'~Spare FB1[273].28'; 8765 '~Spare FB1[273].29'; 8766 '~Spare FB1[273].30'; 8767 '~Spare FB1[273].31'; 8768 '~Spare FB1[274].0'; 8769 '~Spare FB1[274].1'; 8770 '~Spare FB1[274].2'; 8771 '~Spare FB1[274].3'; 8772 '~Spare FB1[274].4'; 8773 '~Spare FB1[274].5'; 8774 '~Spare FB1[274].6'; 8775 '~Spare FB1[274].7'; 8776 '~Spare FB1[274].8'; 8777 '~Spare FB1[274].9'; 8778 '~Spare FB1[274].10'; 8779 '~Spare FB1[274].11'; 8780 '~Spare FB1[274].12'; 8781 '~Spare FB1[274].13'; 8782 '~Spare FB1[274].14'; 8783 '~Spare FB1[274].15'; 8784 '~Spare FB1[274].16'; 8785 '~Spare FB1[274].17'; 8786 '~Spare FB1[274].18'; 8787 '~Spare FB1[274].19'; 8788 '~Spare FB1[274].20'; 8789 '~Spare FB1[274].21'; 8790 '~Spare FB1[274].22'; 8791 '~Spare FB1[274].23'; 8792 '~Spare FB1[274].24'; 8793 '~Spare FB1[274].25'; 8794 '~Spare FB1[274].26'; 8795 '~Spare FB1[274].27'; 8796 '~Spare FB1[274].28'; 8797 '~Spare FB1[274].29'; 8798 '~Spare FB1[274].30'; 8799 '~Spare FB1[274].31'; 8800 '~Spare FB1[275].0'; 8801 '~Spare FB1[275].1'; 8802 '~Spare FB1[275].2'; 8803 '~Spare FB1[275].3'; 8804 '~Spare FB1[275].4'; 8805 '~Spare FB1[275].5'; 8806 '~Spare FB1[275].6'; 8807 '~Spare FB1[275].7'; 8808 '~Spare FB1[275].8'; 8809 '~Spare FB1[275].9'; 8810 '~Spare FB1[275].10'; 8811 '~Spare FB1[275].11'; 8812 '~Spare FB1[275].12'; 8813 '~Spare FB1[275].13'; 8814 '~Spare FB1[275].14'; 8815 '~Spare FB1[275].15'; 8816 '~Spare FB1[275].16'; 8817 '~Spare FB1[275].17'; 8818 '~Spare FB1[275].18'; 8819 '~Spare FB1[275].19'; 8820 '~Spare FB1[275].20'; 8821 '~Spare FB1[275].21'; 8822 '~Spare FB1[275].22'; 8823 '~Spare FB1[275].23'; 8824 '~Spare FB1[275].24'; 8825 '~Spare FB1[275].25'; 8826 '~Spare FB1[275].26'; 8827 '~Spare FB1[275].27'; 8828 '~Spare FB1[275].28'; 8829 '~Spare FB1[275].29'; 8830 '~Spare FB1[275].30'; 8831 '~Spare FB1[275].31'; 8832 '~S001R05CN.I.RbtCtrlFlt - Control Fault FB1[276].0'; 8833 '~S001R05CN.I.CollDetect - Collision Detect FB1[276].1'; 8834 '~S001R05CN.Ix.RbtPromptBox - View Prompt Box at Teach Pendant FB1[276].2'; 8835 '~Spare FB1[276].3'; 8836 '~Spare FB1[276].4'; 8837 '~Spare FB1[276].5'; 8838 '~Spare FB1[276].6'; 8839 '~Spare FB1[276].7'; 8840 '~Spare FB1[276].8'; 8841 '~Spare FB1[276].9'; 8842 '~Spare FB1[276].10'; 8843 '~S001R05CN.I.Wc1WldFlt -Weld Controller 1 Weld Fault FB1[276].11'; 8844 '~S001R05CN.I.Wc1Flt - Weld Timer Flt - Depress Man Weld To Continue FB1[276].12'; 8845 '~S001R05CN.I.Wc1SGunFlt - Weld Controller 1 Servo Gun Fault FB1[276].13'; 8846 '~S001R05CN.I.Wc1SGunMtrTempFlt - Cntrl 1 Servo Gun Motor Over Temp FB1[276].14'; 8847 '~S001R05CN.I.Td1MtrFlt - Tip Dress 1 Motor Fault FB1[276].15'; 8848 '~S001R05CN.I.WC1XfmrTempFlt - Weld Cntrl 1 Transformer Over Temp FB1[276].16'; 8849 '~S001R05CN.I.AutoTipChng1Flt - Auto Tip Changer 1 Fault FB1[276].17'; 8850 '~S001R05CN.I.Slr1NotReady - Seal Controller 1 Not Ready FB1[276].18'; 8851 '~S001R05CN.I.Slr1MajorFlt - Seal Controller 1 Major Fault FB1[276].19'; 8852 '~S001R05CN.I.Slr1VolNotOk - Seal Controller 1 Volume Not Ok Fault FB1[276].20'; 8853 '~S001R05CN.I.Slr1PurgeFlt - Seal Controller 1 Purge Fault FB1[276].21'; 8854 '~S001R05CN.I.Slr1DoserNot Filled - Seal Cntrl 1 Doser Not Filled FB1[276].22'; 8855 '~S001R05CN.I.Slr1No2ClnMxr - Seal Cntrl1 No 2C In Mixer Fault FB1[276].23'; 8856 '~S001R05CN.I.Slr1NzlBroken - Seal Controller 1 Nozzle Broken Fault FB1[276].24'; 8857 '~S001R05CN.I.Slr1NozzleChgReq - Seal Cntrl1 Nozzle Change Reqd FB1[276].25'; 8858 '~S001R05CN.I.Slr1CycleInterrupted - Seal Cntrl1 Cycle Interrupted FB1[276].26'; 8859 '~S001R05CN.I.Stdw1Flt - Stud Weld 1 Weld Fault FB1[276].27'; 8860 '~S001R05CN.I.Stdw1DlyExcdd - Stud Weld 1 Time Delay Exceeded Flt FB1[276].28'; 8861 '~S001R05CN.I.Stdw1Maint Reqd - Stud Weld 1 Maintenance Required FB1[276].29'; 8862 '~S001R05CN.I.Stdw1Reject - Stud Weld 1 art Reject Fault FB1[276].30'; 8863 '~S001R05CN.I.Rvt1Flt - Rivet Controller 1 Fault FB1[276].31'; 8864 '~S001R05CN.I.Rvt1DlyExcdd - Rivet Cntrl 1 Time Delay Exceeded Flt FB1[277].0'; 8865 '~S001R05CN.I.AutoPulledTipByp1 - Auto Pulled Tip Bypass 1 FB1[277].1'; 8866 '~S001R05CN.I.StdWld1EquipmentFlt - Stud Weld 1 Equipment Fault FB1[277].2'; 8867 '~S001R05CN.I.StdWld1BrcktNotPresent - Stud Weld 1 Bracket Not Pres FB1[277].3'; 8868 '~S001R05CN.I.PierceFlt - Pierce Fault FB1[277].4'; 8869 '~S001R05CN.I.NoVisionMeasErr - Vision System Measurement Error FB1[277].5'; 8870 '~S001R05CN.I.VisionSysCalErr - Vision System Calibration Fault FB1[277].6'; 8871 '~S001R05CN.I.VisionSysErr - Vision System Error FB1[277].7'; 8872 '~S001R05CN.I.RackOutOfTolerance - Vision Sys Rack Out Of Tolerance FB1[277].8'; 8873 '~S001R05CN.Ix.TorqFlt - Torque Not Ok FB1[277].9'; 8874 '~S001R05CN.Ix.MwFlt - Mig Weld Controller Fault FB1[277].10'; 8875 '~S001R05CN.Ix.MwWireStuckFlt - Mig Welder Wire Stuck FB1[277].11'; 8876 '~S001R05CN.Ix.MwWldFlt - Mig Welder Bad Bronze Weld Indicator Flt FB1[277].12'; 8877 '~S001R05CN.I.O.TipChngReqd1 - Weld Cntrl 1 Tip Change Required FB1[277].13'; 8878 '~S001R05CN.I.M.NutDetectFlt1 - Nut Welder 1 Nut Detection Fault FB1[277].14'; 8879 '~S001R05CN.I.M.NutProjFlt1 - Nut Welder 1 Weld Not In Tolerance FB1[277].15'; 8880 '~S001R05CN.M.WrongRivetAtNose - Remove Wrong Rivet At Nose FB1[277].16'; 8881 '~S001R05CN.Ix.MwWldLimitErr - Mig Welder CurrentVoltage Out of Tolerance FB1[277].17'; 8882 '~S001R05CN.Ix.MigRdy Mig Welder Not Ready FB1[277].18'; 8883 '~Spare FB1[277].19'; 8884 '~Spare FB1[277].20'; 8885 '~S001R05CN.I.Wc2WldFlt -Weld Controller 2 Weld Fault FB1[277].21'; 8886 '~S001R05CN.I.Wc2Flt - Weld Timer Flt - Depress Man Weld To Continue FB1[277].22'; 8887 '~S001R05CN.I.Wc2SGunFlt - Weld Controller 2 Servo Gun Fault FB1[277].23'; 8888 '~S001R05CN.I.Wc2SGunMtrTempFlt - Cntrl 2 Servo Gun Motor Over Temp FB1[277].24'; 8889 '~S001R05CN.I.Td2MtrFlt - Tip Dress 2 Motor Fault FB1[277].25'; 8890 '~S001R05CN.I.WC2XfmrTempFlt - Weld Cntrl 2 Transformer Over Temp FB1[277].26'; 8891 '~S001R05CN.I.AutoTipChng2Flt - Auto Tip Changer 2 Fault FB1[277].27'; 8892 '~S001R05CN.I.Slr2NotReady - Seal Controller 2 Not Ready FB1[277].28'; 8893 '~S001R05CN.I.Slr2MajorFlt - Seal Controller 2 Major Fault FB1[277].29'; 8894 '~S001R05CN.I.Slr2VolNotOk - Seal Controller 2 Volume Not Ok Fault FB1[277].30'; 8895 '~S001R05CN.I.Slr2PurgeFlt - Seal Controller 2 Purge Fault FB1[277].31'; 8896 '~S001R05CN.I.Slr2DoserNot Filled - Seal Cntrl 2 Doser Not Filled FB1[278].0'; 8897 '~S001R05CN.I.Slr2No2ClnMxr - Seal Cntrl2 No 2C In Mixer Fault FB1[278].1'; 8898 '~S001R05CN.I.Slr2NzlBroken - Seal Controller 2 Nozzle Broken Fault FB1[278].2'; 8899 '~S001R05CN.I.Slr2NozzleChgReq - Seal Cntrl2 Nozzle Change Reqd FB1[278].3'; 8900 '~S001R05CN.I.Slr2CycleInterrupted - Seal Cntrl2 Cycle Interrupted FB1[278].4'; 8901 '~S001R05CN.I.Stdw2Flt - Stud Weld 2 Weld Fault FB1[278].5'; 8902 '~S001R05CN.I.Stdw2DlyExcdd - Stud Weld 2 Time Delay Exceeded Flt FB1[278].6'; 8903 '~S001R05CN.I.Stdw2Maint Reqd - Stud Weld 2 Maintenance Required FB1[278].7'; 8904 '~S001R05CN.I.Stdw2Reject - Stud Weld 2 art Reject Fault FB1[278].8'; 8905 '~S001R05CN.I.Rvt2Flt - Rivet Controller 2 Fault FB1[278].9'; 8906 '~S001R05CN.I.Rvt2DlyExcdd - Rivet Cntrl 2 Time Delay Exceeded Flt FB1[278].10'; 8907 '~S001R05CN.I.AutoPulledTipByp2 - Auto Pulled Tip Bypass 2 FB1[278].11'; 8908 '~S001R05CN.I.StdWld2EquipmentFlt - Stud Weld 2 Equipment Fault FB1[278].12'; 8909 '~S001R05CN.I.StdWld2BrcktNotPresent - Stud Weld 2 Bracket Not Pres FB1[278].13'; 8910 '~S001R05CN.Ix.LsrWldMntrFlt - Seam Geometry/Laser Weld Monitor Flt FB1[278].14'; 8911 '~S001R05CN.Ix.LsrHeadFlt - Laser Head Fault FB1[278].15'; 8912 '~S001R05CN.Ix.LsrGlsFlt - Glass Fault FB1[278].16'; 8913 '~S001R05CN.Ix.LsrWhlFlt - Pressure Wheel Not In Range Fault FB1[278].17'; 8914 '~S001R05CN.Ix.LsrGeoFlt - Seam Geometry/Laser Bad Process Geo Flt FB1[278].18'; 8915 '~S001R05CN.Ix.LsrHdCollFlt - Laser Head Collision Fault FB1[278].19'; 8916 '~S001R05CN.Ix.LsrHdSysFlt - Laser Head System Fault FB1[278].20'; 8917 '~S001R05CN.Ix.LsrHdFar - Laser Head Far Fault FB1[278].21'; 8918 '~S001R05CN.Ix.LsrHdSftCollFlt - Laser Head Software Collision Flt FB1[278].22'; 8919 '~S001R05CN.I.O.TipChngReqd2 - Weld Cntrl 2 Tip Change Required FB1[278].23'; 8920 '~S001R05CN.I.M.NutDetectFlt2 - Nut Welder 2 Nut Detection Fault FB1[278].24'; 8921 '~S001R05CN.I.M.NutProjFlt2 - Nut Welder 2 Weld Not In Tolerance FB1[278].25'; 8922 '~S001R05CN.I.TCWrongToolInStand - Tool Changer Wrong Tool In Stand FB1[278].26'; 8923 '~Spare FB1[278].27'; 8924 '~Spare FB1[278].28'; 8925 '~Spare FB1[278].29'; 8926 '~Spare FB1[278].30'; 8927 '~Spare FB1[278].31'; 8928 '~S001R05CN.I.VisionCommOK - Vision System Comm Fault FB1[279].0'; 8929 '~S001R05CN.I.OutOfTolerance - Vision System Out Of Tolerance FB1[279].1'; 8930 '~S001R05CN.I.MeasureReject - Vision System Measure Reject FB1[279].2'; 8931 '~S001R05CN.I.VisionSysCalibrationFlt - Vision System Calibration Flt FB1[279].3'; 8932 '~S001R05CN.I.VisionSysFlt - Vision System Flt FB1[279].4'; 8933 '~Spare FB1[279].5'; 8934 '~Spare FB1[279].6'; 8935 '~Spare FB1[279].7'; 8936 '~Spare FB1[279].8'; 8937 '~Spare FB1[279].9'; 8938 '~Spare FB1[279].10'; 8939 '~Spare FB1[279].11'; 8940 '~Spare FB1[279].12'; 8941 '~Spare FB1[279].13'; 8942 '~Spare FB1[279].14'; 8943 '~Spare FB1[279].15'; 8944 '~Spare FB1[279].16'; 8945 '~Spare FB1[279].17'; 8946 '~S001R05CN.M.InteruptCyc - Laser Cyc Interupt Cut Wire And Reject Car FB1[279].18'; 8947 '~S001R05CN.M.SuspectPart Inspect Vehicle And Accept Or Reject FB1[279].19'; 8948 '~S001R05 Power Meter High Power Fault Detected FB1[279].20'; 8949 '~S001R05 Power Meter Low Power Fault Detected FB1[279].21'; 8950 '~Spare FB1[279].22'; 8951 '~Spare FB1[279].23'; 8952 '~Spare FB1[279].24'; 8953 '~Spare FB1[279].25'; 8954 '~Spare FB1[279].26'; 8955 '~Spare FB1[279].27'; 8956 '~Spare FB1[279].28'; 8957 '~Spare FB1[279].29'; 8958 '~Spare FB1[279].30'; 8959 '~Spare FB1[279].31'; 8960 '~Spare FB1[280].0'; 8961 '~Spare FB1[280].1'; 8962 '~Spare FB1[280].2'; 8963 '~Spare FB1[280].3'; 8964 '~Spare FB1[280].4'; 8965 '~Spare FB1[280].5'; 8966 '~Spare FB1[280].6'; 8967 '~Spare FB1[280].7'; 8968 '~Spare FB1[280].8'; 8969 '~Spare FB1[280].9'; 8970 '~Spare FB1[280].10'; 8971 '~Spare FB1[280].11'; 8972 '~Spare FB1[280].12'; 8973 '~Spare FB1[280].13'; 8974 '~Spare FB1[280].14'; 8975 '~Spare FB1[280].15'; 8976 '~Spare FB1[280].16'; 8977 '~Spare FB1[280].17'; 8978 '~Spare FB1[280].18'; 8979 '~Spare FB1[280].19'; 8980 '~Spare FB1[280].20'; 8981 '~Spare FB1[280].21'; 8982 '~Spare FB1[280].22'; 8983 '~Spare FB1[280].23'; 8984 '~Spare FB1[280].24'; 8985 '~Spare FB1[280].25'; 8986 '~Spare FB1[280].26'; 8987 '~Spare FB1[280].27'; 8988 '~Spare FB1[280].28'; 8989 '~Spare FB1[280].29'; 8990 '~Spare FB1[280].30'; 8991 '~Spare FB1[280].31'; 8992 '~Spare FB1[281].0'; 8993 '~Spare FB1[281].1'; 8994 '~Spare FB1[281].2'; 8995 '~Spare FB1[281].3'; 8996 '~Spare FB1[281].4'; 8997 '~Spare FB1[281].5'; 8998 '~Spare FB1[281].6'; 8999 '~Spare FB1[281].7'; 9000 '~Spare FB1[281].8'; 9001 '~Spare FB1[281].9'; 9002 '~Spare FB1[281].10'; 9003 '~Spare FB1[281].11'; 9004 '~Spare FB1[281].12'; 9005 '~Spare FB1[281].13'; 9006 '~Spare FB1[281].14'; 9007 '~Spare FB1[281].15'; 9008 '~Spare FB1[281].16'; 9009 '~Spare FB1[281].17'; 9010 '~Spare FB1[281].18'; 9011 '~Spare FB1[281].19'; 9012 '~Spare FB1[281].20'; 9013 '~Spare FB1[281].21'; 9014 '~Spare FB1[281].22'; 9015 '~Spare FB1[281].23'; 9016 '~Spare FB1[281].24'; 9017 '~Spare FB1[281].25'; 9018 '~Spare FB1[281].26'; 9019 '~Spare FB1[281].27'; 9020 '~Spare FB1[281].28'; 9021 '~Spare FB1[281].29'; 9022 '~Spare FB1[281].30'; 9023 '~Spare FB1[281].31'; 9024 '~Spare FB1[282].0'; 9025 '~Spare FB1[282].1'; 9026 '~Spare FB1[282].2'; 9027 '~Spare FB1[282].3'; 9028 '~Spare FB1[282].4'; 9029 '~Spare FB1[282].5'; 9030 '~Spare FB1[282].6'; 9031 '~Spare FB1[282].7'; 9032 '~Spare FB1[282].8'; 9033 '~Spare FB1[282].9'; 9034 '~Spare FB1[282].10'; 9035 '~Spare FB1[282].11'; 9036 '~Spare FB1[282].12'; 9037 '~Spare FB1[282].13'; 9038 '~Spare FB1[282].14'; 9039 '~Spare FB1[282].15'; 9040 '~Spare FB1[282].16'; 9041 '~Spare FB1[282].17'; 9042 '~Spare FB1[282].18'; 9043 '~Spare FB1[282].19'; 9044 '~Spare FB1[282].20'; 9045 '~Spare FB1[282].21'; 9046 '~Spare FB1[282].22'; 9047 '~Spare FB1[282].23'; 9048 '~Spare FB1[282].24'; 9049 '~Spare FB1[282].25'; 9050 '~Spare FB1[282].26'; 9051 '~Spare FB1[282].27'; 9052 '~Spare FB1[282].28'; 9053 '~Spare FB1[282].29'; 9054 '~Spare FB1[282].30'; 9055 '~Spare FB1[282].31'; 9056 '~Spare FB1[283].0'; 9057 '~Spare FB1[283].1'; 9058 '~Spare FB1[283].2'; 9059 '~Spare FB1[283].3'; 9060 '~Spare FB1[283].4'; 9061 '~Spare FB1[283].5'; 9062 '~Spare FB1[283].6'; 9063 '~Spare FB1[283].7'; 9064 '~Spare FB1[283].8'; 9065 '~Spare FB1[283].9'; 9066 '~Spare FB1[283].10'; 9067 '~Spare FB1[283].11'; 9068 '~Spare FB1[283].12'; 9069 '~Spare FB1[283].13'; 9070 '~Spare FB1[283].14'; 9071 '~Spare FB1[283].15'; 9072 '~Spare FB1[283].16'; 9073 '~Spare FB1[283].17'; 9074 '~Spare FB1[283].18'; 9075 '~Spare FB1[283].19'; 9076 '~Spare FB1[283].20'; 9077 '~Spare FB1[283].21'; 9078 '~Spare FB1[283].22'; 9079 '~Spare FB1[283].23'; 9080 '~Spare FB1[283].24'; 9081 '~Spare FB1[283].25'; 9082 '~Spare FB1[283].26'; 9083 '~Spare FB1[283].27'; 9084 '~Spare FB1[283].28'; 9085 '~Spare FB1[283].29'; 9086 '~Spare FB1[283].30'; 9087 '~Spare FB1[283].31'; 9088 '~S001R06CN.I.RbtCtrlFlt - Control Fault FB1[284].0'; 9089 '~S001R06CN.I.CollDetect - Collision Detect FB1[284].1'; 9090 '~S001R06CN.Ix.RbtPromptBox - View Prompt Box at Teach Pendant FB1[284].2'; 9091 '~Spare FB1[284].3'; 9092 '~Spare FB1[284].4'; 9093 '~Spare FB1[284].5'; 9094 '~Spare FB1[284].6'; 9095 '~Spare FB1[284].7'; 9096 '~Spare FB1[284].8'; 9097 '~Spare FB1[284].9'; 9098 '~Spare FB1[284].10'; 9099 '~S001R06CN.I.Wc1WldFlt -Weld Controller 1 Weld Fault FB1[284].11'; 9100 '~S001R06CN.I.Wc1Flt - Weld Timer Flt - Depress Man Weld To Continue FB1[284].12'; 9101 '~S001R06CN.I.Wc1SGunFlt - Weld Controller 1 Servo Gun Fault FB1[284].13'; 9102 '~S001R06CN.I.Wc1SGunMtrTempFlt - Cntrl 1 Servo Gun Motor Over Temp FB1[284].14'; 9103 '~S001R06CN.I.Td1MtrFlt - Tip Dress 1 Motor Fault FB1[284].15'; 9104 '~S001R06CN.I.WC1XfmrTempFlt - Weld Cntrl 1 Transformer Over Temp FB1[284].16'; 9105 '~S001R06CN.I.AutoTipChng1Flt - Auto Tip Changer 1 Fault FB1[284].17'; 9106 '~S001R06CN.I.Slr1NotReady - Seal Controller 1 Not Ready FB1[284].18'; 9107 '~S001R06CN.I.Slr1MajorFlt - Seal Controller 1 Major Fault FB1[284].19'; 9108 '~S001R06CN.I.Slr1VolNotOk - Seal Controller 1 Volume Not Ok Fault FB1[284].20'; 9109 '~S001R06CN.I.Slr1PurgeFlt - Seal Controller 1 Purge Fault FB1[284].21'; 9110 '~S001R06CN.I.Slr1DoserNot Filled - Seal Cntrl 1 Doser Not Filled FB1[284].22'; 9111 '~S001R06CN.I.Slr1No2ClnMxr - Seal Cntrl1 No 2C In Mixer Fault FB1[284].23'; 9112 '~S001R06CN.I.Slr1NzlBroken - Seal Controller 1 Nozzle Broken Fault FB1[284].24'; 9113 '~S001R06CN.I.Slr1NozzleChgReq - Seal Cntrl1 Nozzle Change Reqd FB1[284].25'; 9114 '~S001R06CN.I.Slr1CycleInterrupted - Seal Cntrl1 Cycle Interrupted FB1[284].26'; 9115 '~S001R06CN.I.Stdw1Flt - Stud Weld 1 Weld Fault FB1[284].27'; 9116 '~S001R06CN.I.Stdw1DlyExcdd - Stud Weld 1 Time Delay Exceeded Flt FB1[284].28'; 9117 '~S001R06CN.I.Stdw1Maint Reqd - Stud Weld 1 Maintenance Required FB1[284].29'; 9118 '~S001R06CN.I.Stdw1Reject - Stud Weld 1 art Reject Fault FB1[284].30'; 9119 '~S001R06CN.I.Rvt1Flt - Rivet Controller 1 Fault FB1[284].31'; 9120 '~S001R06CN.I.Rvt1DlyExcdd - Rivet Cntrl 1 Time Delay Exceeded Flt FB1[285].0'; 9121 '~S001R06CN.I.AutoPulledTipByp1 - Auto Pulled Tip Bypass 1 FB1[285].1'; 9122 '~S001R06CN.I.StdWld1EquipmentFlt - Stud Weld 1 Equipment Fault FB1[285].2'; 9123 '~S001R06CN.I.StdWld1BrcktNotPresent - Stud Weld 1 Bracket Not Pres FB1[285].3'; 9124 '~S001R06CN.I.PierceFlt - Pierce Fault FB1[285].4'; 9125 '~S001R06CN.I.NoVisionMeasErr - Vision System Measurement Error FB1[285].5'; 9126 '~S001R06CN.I.VisionSysCalErr - Vision System Calibration Fault FB1[285].6'; 9127 '~S001R06CN.I.VisionSysErr - Vision System Error FB1[285].7'; 9128 '~S001R06CN.I.RackOutOfTolerance - Vision Sys Rack Out Of Tolerance FB1[285].8'; 9129 '~S001R06CN.Ix.TorqFlt - Torque Not Ok FB1[285].9'; 9130 '~S001R06CN.Ix.MwFlt - Mig Weld Controller Fault FB1[285].10'; 9131 '~S001R06CN.Ix.MwWireStuckFlt - Mig Welder Wire Stuck FB1[285].11'; 9132 '~S001R06CN.Ix.MwWldFlt - Mig Welder Bad Bronze Weld Indicator Flt FB1[285].12'; 9133 '~S001R06CN.I.O.TipChngReqd1 - Weld Cntrl 1 Tip Change Required FB1[285].13'; 9134 '~S001R06CN.I.M.NutDetectFlt1 - Nut Welder 1 Nut Detection Fault FB1[285].14'; 9135 '~S001R06CN.I.M.NutProjFlt1 - Nut Welder 1 Weld Not In Tolerance FB1[285].15'; 9136 '~S001R06CN.M.WrongRivetAtNose - Remove Wrong Rivet At Nose FB1[285].16'; 9137 '~S001R06CN.Ix.MwWldLimitErr - Mig Welder CurrentVoltage Out of Tolerance FB1[285].17'; 9138 '~S001R06CN.Ix.MigRdy Mig Welder Not Ready FB1[285].18'; 9139 '~Spare FB1[285].19'; 9140 '~Spare FB1[285].20'; 9141 '~S001R06CN.I.Wc2WldFlt -Weld Controller 2 Weld Fault FB1[285].21'; 9142 '~S001R06CN.I.Wc2Flt - Weld Timer Flt - Depress Man Weld To Continue FB1[285].22'; 9143 '~S001R06CN.I.Wc2SGunFlt - Weld Controller 2 Servo Gun Fault FB1[285].23'; 9144 '~S001R06CN.I.Wc2SGunMtrTempFlt - Cntrl 2 Servo Gun Motor Over Temp FB1[285].24'; 9145 '~S001R06CN.I.Td2MtrFlt - Tip Dress 2 Motor Fault FB1[285].25'; 9146 '~S001R06CN.I.WC2XfmrTempFlt - Weld Cntrl 2 Transformer Over Temp FB1[285].26'; 9147 '~S001R06CN.I.AutoTipChng2Flt - Auto Tip Changer 2 Fault FB1[285].27'; 9148 '~S001R06CN.I.Slr2NotReady - Seal Controller 2 Not Ready FB1[285].28'; 9149 '~S001R06CN.I.Slr2MajorFlt - Seal Controller 2 Major Fault FB1[285].29'; 9150 '~S001R06CN.I.Slr2VolNotOk - Seal Controller 2 Volume Not Ok Fault FB1[285].30'; 9151 '~S001R06CN.I.Slr2PurgeFlt - Seal Controller 2 Purge Fault FB1[285].31'; 9152 '~S001R06CN.I.Slr2DoserNot Filled - Seal Cntrl 2 Doser Not Filled FB1[286].0'; 9153 '~S001R06CN.I.Slr2No2ClnMxr - Seal Cntrl2 No 2C In Mixer Fault FB1[286].1'; 9154 '~S001R06CN.I.Slr2NzlBroken - Seal Controller 2 Nozzle Broken Fault FB1[286].2'; 9155 '~S001R06CN.I.Slr2NozzleChgReq - Seal Cntrl2 Nozzle Change Reqd FB1[286].3'; 9156 '~S001R06CN.I.Slr2CycleInterrupted - Seal Cntrl2 Cycle Interrupted FB1[286].4'; 9157 '~S001R06CN.I.Stdw2Flt - Stud Weld 2 Weld Fault FB1[286].5'; 9158 '~S001R06CN.I.Stdw2DlyExcdd - Stud Weld 2 Time Delay Exceeded Flt FB1[286].6'; 9159 '~S001R06CN.I.Stdw2Maint Reqd - Stud Weld 2 Maintenance Required FB1[286].7'; 9160 '~S001R06CN.I.Stdw2Reject - Stud Weld 2 art Reject Fault FB1[286].8'; 9161 '~S001R06CN.I.Rvt2Flt - Rivet Controller 2 Fault FB1[286].9'; 9162 '~S001R06CN.I.Rvt2DlyExcdd - Rivet Cntrl 2 Time Delay Exceeded Flt FB1[286].10'; 9163 '~S001R06CN.I.AutoPulledTipByp2 - Auto Pulled Tip Bypass 2 FB1[286].11'; 9164 '~S001R06CN.I.StdWld2EquipmentFlt - Stud Weld 2 Equipment Fault FB1[286].12'; 9165 '~S001R06CN.I.StdWld2BrcktNotPresent - Stud Weld 2 Bracket Not Pres FB1[286].13'; 9166 '~S001R06CN.Ix.LsrWldMntrFlt - Seam Geometry/Laser Weld Monitor Flt FB1[286].14'; 9167 '~S001R06CN.Ix.LsrHeadFlt - Laser Head Fault FB1[286].15'; 9168 '~S001R06CN.Ix.LsrGlsFlt - Glass Fault FB1[286].16'; 9169 '~S001R06CN.Ix.LsrWhlFlt - Pressure Wheel Not In Range Fault FB1[286].17'; 9170 '~S001R06CN.Ix.LsrGeoFlt - Seam Geometry/Laser Bad Process Geo Flt FB1[286].18'; 9171 '~S001R06CN.Ix.LsrHdCollFlt - Laser Head Collision Fault FB1[286].19'; 9172 '~S001R06CN.Ix.LsrHdSysFlt - Laser Head System Fault FB1[286].20'; 9173 '~S001R06CN.Ix.LsrHdFar - Laser Head Far Fault FB1[286].21'; 9174 '~S001R06CN.Ix.LsrHdSftCollFlt - Laser Head Software Collision Flt FB1[286].22'; 9175 '~S001R06CN.I.O.TipChngReqd2 - Weld Cntrl 2 Tip Change Required FB1[286].23'; 9176 '~S001R06CN.I.M.NutDetectFlt2 - Nut Welder 2 Nut Detection Fault FB1[286].24'; 9177 '~S001R06CN.I.M.NutProjFlt2 - Nut Welder 2 Weld Not In Tolerance FB1[286].25'; 9178 '~S001R06CN.I.TCWrongToolInStand - Tool Changer Wrong Tool In Stand FB1[286].26'; 9179 '~Spare FB1[286].27'; 9180 '~Spare FB1[286].28'; 9181 '~Spare FB1[286].29'; 9182 '~Spare FB1[286].30'; 9183 '~Spare FB1[286].31'; 9184 '~S001R06CN.I.VisionCommOK - Vision System Comm Fault FB1[287].0'; 9185 '~S001R06CN.I.OutOfTolerance - Vision System Out Of Tolerance FB1[287].1'; 9186 '~S001R06CN.I.MeasureReject - Vision System Measure Reject FB1[287].2'; 9187 '~S001R06CN.I.VisionSysCalibrationFlt - Vision System Calibration Flt FB1[287].3'; 9188 '~S001R06CN.I.VisionSysFlt - Vision System Flt FB1[287].4'; 9189 '~Spare FB1[287].5'; 9190 '~Spare FB1[287].6'; 9191 '~Spare FB1[287].7'; 9192 '~Spare FB1[287].8'; 9193 '~Spare FB1[287].9'; 9194 '~Spare FB1[287].10'; 9195 '~Spare FB1[287].11'; 9196 '~Spare FB1[287].12'; 9197 '~Spare FB1[287].13'; 9198 '~Spare FB1[287].14'; 9199 '~Spare FB1[287].15'; 9200 '~Spare FB1[287].16'; 9201 '~Spare FB1[287].17'; 9202 '~S001R06CN.M.InteruptCyc - Laser Cyc Interupt Cut Wire And Reject Car FB1[287].18'; 9203 '~S001R06CN.M.SuspectPart Inspect Vehicle And Accept Or Reject FB1[287].19'; 9204 '~S001R06 Power Meter High Power Fault Detected FB1[287].20'; 9205 '~S001R06 Power Meter Low Power Fault Detected FB1[287].21'; 9206 '~Spare FB1[287].22'; 9207 '~Spare FB1[287].23'; 9208 '~Spare FB1[287].24'; 9209 '~Spare FB1[287].25'; 9210 '~Spare FB1[287].26'; 9211 '~Spare FB1[287].27'; 9212 '~Spare FB1[287].28'; 9213 '~Spare FB1[287].29'; 9214 '~Spare FB1[287].30'; 9215 '~Spare FB1[287].31'; 9216 '~Spare FB1[288].0'; 9217 '~Spare FB1[288].1'; 9218 '~Spare FB1[288].2'; 9219 '~Spare FB1[288].3'; 9220 '~Spare FB1[288].4'; 9221 '~Spare FB1[288].5'; 9222 '~Spare FB1[288].6'; 9223 '~Spare FB1[288].7'; 9224 '~Spare FB1[288].8'; 9225 '~Spare FB1[288].9'; 9226 '~Spare FB1[288].10'; 9227 '~Spare FB1[288].11'; 9228 '~Spare FB1[288].12'; 9229 '~Spare FB1[288].13'; 9230 '~Spare FB1[288].14'; 9231 '~Spare FB1[288].15'; 9232 '~Spare FB1[288].16'; 9233 '~Spare FB1[288].17'; 9234 '~Spare FB1[288].18'; 9235 '~Spare FB1[288].19'; 9236 '~Spare FB1[288].20'; 9237 '~Spare FB1[288].21'; 9238 '~Spare FB1[288].22'; 9239 '~Spare FB1[288].23'; 9240 '~Spare FB1[288].24'; 9241 '~Spare FB1[288].25'; 9242 '~Spare FB1[288].26'; 9243 '~Spare FB1[288].27'; 9244 '~Spare FB1[288].28'; 9245 '~Spare FB1[288].29'; 9246 '~Spare FB1[288].30'; 9247 '~Spare FB1[288].31'; 9248 '~Spare FB1[289].0'; 9249 '~Spare FB1[289].1'; 9250 '~Spare FB1[289].2'; 9251 '~Spare FB1[289].3'; 9252 '~Spare FB1[289].4'; 9253 '~Spare FB1[289].5'; 9254 '~Spare FB1[289].6'; 9255 '~Spare FB1[289].7'; 9256 '~Spare FB1[289].8'; 9257 '~Spare FB1[289].9'; 9258 '~Spare FB1[289].10'; 9259 '~Spare FB1[289].11'; 9260 '~Spare FB1[289].12'; 9261 '~Spare FB1[289].13'; 9262 '~Spare FB1[289].14'; 9263 '~Spare FB1[289].15'; 9264 '~Spare FB1[289].16'; 9265 '~Spare FB1[289].17'; 9266 '~Spare FB1[289].18'; 9267 '~Spare FB1[289].19'; 9268 '~Spare FB1[289].20'; 9269 '~Spare FB1[289].21'; 9270 '~Spare FB1[289].22'; 9271 '~Spare FB1[289].23'; 9272 '~Spare FB1[289].24'; 9273 '~Spare FB1[289].25'; 9274 '~Spare FB1[289].26'; 9275 '~Spare FB1[289].27'; 9276 '~Spare FB1[289].28'; 9277 '~Spare FB1[289].29'; 9278 '~Spare FB1[289].30'; 9279 '~Spare FB1[289].31'; 9280 '~Spare FB1[290].0'; 9281 '~Spare FB1[290].1'; 9282 '~Spare FB1[290].2'; 9283 '~Spare FB1[290].3'; 9284 '~Spare FB1[290].4'; 9285 '~Spare FB1[290].5'; 9286 '~Spare FB1[290].6'; 9287 '~Spare FB1[290].7'; 9288 '~Spare FB1[290].8'; 9289 '~Spare FB1[290].9'; 9290 '~Spare FB1[290].10'; 9291 '~Spare FB1[290].11'; 9292 '~Spare FB1[290].12'; 9293 '~Spare FB1[290].13'; 9294 '~Spare FB1[290].14'; 9295 '~Spare FB1[290].15'; 9296 '~Spare FB1[290].16'; 9297 '~Spare FB1[290].17'; 9298 '~Spare FB1[290].18'; 9299 '~Spare FB1[290].19'; 9300 '~Spare FB1[290].20'; 9301 '~Spare FB1[290].21'; 9302 '~Spare FB1[290].22'; 9303 '~Spare FB1[290].23'; 9304 '~Spare FB1[290].24'; 9305 '~Spare FB1[290].25'; 9306 '~Spare FB1[290].26'; 9307 '~Spare FB1[290].27'; 9308 '~Spare FB1[290].28'; 9309 '~Spare FB1[290].29'; 9310 '~Spare FB1[290].30'; 9311 '~Spare FB1[290].31'; 9312 '~Spare FB1[291].0'; 9313 '~Spare FB1[291].1'; 9314 '~Spare FB1[291].2'; 9315 '~Spare FB1[291].3'; 9316 '~Spare FB1[291].4'; 9317 '~Spare FB1[291].5'; 9318 '~Spare FB1[291].6'; 9319 '~Spare FB1[291].7'; 9320 '~Spare FB1[291].8'; 9321 '~Spare FB1[291].9'; 9322 '~Spare FB1[291].10'; 9323 '~Spare FB1[291].11'; 9324 '~Spare FB1[291].12'; 9325 '~Spare FB1[291].13'; 9326 '~Spare FB1[291].14'; 9327 '~Spare FB1[291].15'; 9328 '~Spare FB1[291].16'; 9329 '~Spare FB1[291].17'; 9330 '~Spare FB1[291].18'; 9331 '~Spare FB1[291].19'; 9332 '~Spare FB1[291].20'; 9333 '~Spare FB1[291].21'; 9334 '~Spare FB1[291].22'; 9335 '~Spare FB1[291].23'; 9336 '~Spare FB1[291].24'; 9337 '~Spare FB1[291].25'; 9338 '~Spare FB1[291].26'; 9339 '~Spare FB1[291].27'; 9340 '~Spare FB1[291].28'; 9341 '~Spare FB1[291].29'; 9342 '~Spare FB1[291].30'; 9343 '~Spare FB1[291].31'; 9344 '~S001R07CN.I.RbtCtrlFlt - Control Fault FB1[292].0'; 9345 '~S001R07CN.I.CollDetect - Collision Detect FB1[292].1'; 9346 '~S001R07CN.Ix.RbtPromptBox - View Prompt Box at Teach Pendant FB1[292].2'; 9347 '~Spare FB1[292].3'; 9348 '~Spare FB1[292].4'; 9349 '~Spare FB1[292].5'; 9350 '~Spare FB1[292].6'; 9351 '~Spare FB1[292].7'; 9352 '~Spare FB1[292].8'; 9353 '~Spare FB1[292].9'; 9354 '~Spare FB1[292].10'; 9355 '~S001R07CN.I.Wc1WldFlt -Weld Controller 1 Weld Fault FB1[292].11'; 9356 '~S001R07CN.I.Wc1Flt - Weld Timer Flt - Depress Man Weld To Continue FB1[292].12'; 9357 '~S001R07CN.I.Wc1SGunFlt - Weld Controller 1 Servo Gun Fault FB1[292].13'; 9358 '~S001R07CN.I.Wc1SGunMtrTempFlt - Cntrl 1 Servo Gun Motor Over Temp FB1[292].14'; 9359 '~S001R07CN.I.Td1MtrFlt - Tip Dress 1 Motor Fault FB1[292].15'; 9360 '~S001R07CN.I.WC1XfmrTempFlt - Weld Cntrl 1 Transformer Over Temp FB1[292].16'; 9361 '~S001R07CN.I.AutoTipChng1Flt - Auto Tip Changer 1 Fault FB1[292].17'; 9362 '~S001R07CN.I.Slr1NotReady - Seal Controller 1 Not Ready FB1[292].18'; 9363 '~S001R07CN.I.Slr1MajorFlt - Seal Controller 1 Major Fault FB1[292].19'; 9364 '~S001R07CN.I.Slr1VolNotOk - Seal Controller 1 Volume Not Ok Fault FB1[292].20'; 9365 '~S001R07CN.I.Slr1PurgeFlt - Seal Controller 1 Purge Fault FB1[292].21'; 9366 '~S001R07CN.I.Slr1DoserNot Filled - Seal Cntrl 1 Doser Not Filled FB1[292].22'; 9367 '~S001R07CN.I.Slr1No2ClnMxr - Seal Cntrl1 No 2C In Mixer Fault FB1[292].23'; 9368 '~S001R07CN.I.Slr1NzlBroken - Seal Controller 1 Nozzle Broken Fault FB1[292].24'; 9369 '~S001R07CN.I.Slr1NozzleChgReq - Seal Cntrl1 Nozzle Change Reqd FB1[292].25'; 9370 '~S001R07CN.I.Slr1CycleInterrupted - Seal Cntrl1 Cycle Interrupted FB1[292].26'; 9371 '~S001R07CN.I.Stdw1Flt - Stud Weld 1 Weld Fault FB1[292].27'; 9372 '~S001R07CN.I.Stdw1DlyExcdd - Stud Weld 1 Time Delay Exceeded Flt FB1[292].28'; 9373 '~S001R07CN.I.Stdw1Maint Reqd - Stud Weld 1 Maintenance Required FB1[292].29'; 9374 '~S001R07CN.I.Stdw1Reject - Stud Weld 1 art Reject Fault FB1[292].30'; 9375 '~S001R07CN.I.Rvt1Flt - Rivet Controller 1 Fault FB1[292].31'; 9376 '~S001R07CN.I.Rvt1DlyExcdd - Rivet Cntrl 1 Time Delay Exceeded Flt FB1[293].0'; 9377 '~S001R07CN.I.AutoPulledTipByp1 - Auto Pulled Tip Bypass 1 FB1[293].1'; 9378 '~S001R07CN.I.StdWld1EquipmentFlt - Stud Weld 1 Equipment Fault FB1[293].2'; 9379 '~S001R07CN.I.StdWld1BrcktNotPresent - Stud Weld 1 Bracket Not Pres FB1[293].3'; 9380 '~S001R07CN.I.PierceFlt - Pierce Fault FB1[293].4'; 9381 '~S001R07CN.I.NoVisionMeasErr - Vision System Measurement Error FB1[293].5'; 9382 '~S001R07CN.I.VisionSysCalErr - Vision System Calibration Fault FB1[293].6'; 9383 '~S001R07CN.I.VisionSysErr - Vision System Error FB1[293].7'; 9384 '~S001R07CN.I.RackOutOfTolerance - Vision Sys Rack Out Of Tolerance FB1[293].8'; 9385 '~S001R07CN.Ix.TorqFlt - Torque Not Ok FB1[293].9'; 9386 '~S001R07CN.Ix.MwFlt - Mig Weld Controller Fault FB1[293].10'; 9387 '~S001R07CN.Ix.MwWireStuckFlt - Mig Welder Wire Stuck FB1[293].11'; 9388 '~S001R07CN.Ix.MwWldFlt - Mig Welder Bad Bronze Weld Indicator Flt FB1[293].12'; 9389 '~S001R07CN.I.O.TipChngReqd1 - Weld Cntrl 1 Tip Change Required FB1[293].13'; 9390 '~S001R07CN.I.M.NutDetectFlt1 - Nut Welder 1 Nut Detection Fault FB1[293].14'; 9391 '~S001R07CN.I.M.NutProjFlt1 - Nut Welder 1 Weld Not In Tolerance FB1[293].15'; 9392 '~S001R07CN.M.WrongRivetAtNose - Remove Wrong Rivet At Nose FB1[293].16'; 9393 '~S001R07CN.Ix.MwWldLimitErr - Mig Welder CurrentVoltage Out of Tolerance FB1[293].17'; 9394 '~S001R07CN.Ix.MigRdy Mig Welder Not Ready FB1[293].18'; 9395 '~Spare FB1[293].19'; 9396 '~Spare FB1[293].20'; 9397 '~S001R07CN.I.Wc2WldFlt -Weld Controller 2 Weld Fault FB1[293].21'; 9398 '~S001R07CN.I.Wc2Flt - Weld Timer Flt - Depress Man Weld To Continue FB1[293].22'; 9399 '~S001R07CN.I.Wc2SGunFlt - Weld Controller 2 Servo Gun Fault FB1[293].23'; 9400 '~S001R07CN.I.Wc2SGunMtrTempFlt - Cntrl 2 Servo Gun Motor Over Temp FB1[293].24'; 9401 '~S001R07CN.I.Td2MtrFlt - Tip Dress 2 Motor Fault FB1[293].25'; 9402 '~S001R07CN.I.WC2XfmrTempFlt - Weld Cntrl 2 Transformer Over Temp FB1[293].26'; 9403 '~S001R07CN.I.AutoTipChng2Flt - Auto Tip Changer 2 Fault FB1[293].27'; 9404 '~S001R07CN.I.Slr2NotReady - Seal Controller 2 Not Ready FB1[293].28'; 9405 '~S001R07CN.I.Slr2MajorFlt - Seal Controller 2 Major Fault FB1[293].29'; 9406 '~S001R07CN.I.Slr2VolNotOk - Seal Controller 2 Volume Not Ok Fault FB1[293].30'; 9407 '~S001R07CN.I.Slr2PurgeFlt - Seal Controller 2 Purge Fault FB1[293].31'; 9408 '~S001R07CN.I.Slr2DoserNot Filled - Seal Cntrl 2 Doser Not Filled FB1[294].0'; 9409 '~S001R07CN.I.Slr2No2ClnMxr - Seal Cntrl2 No 2C In Mixer Fault FB1[294].1'; 9410 '~S001R07CN.I.Slr2NzlBroken - Seal Controller 2 Nozzle Broken Fault FB1[294].2'; 9411 '~S001R07CN.I.Slr2NozzleChgReq - Seal Cntrl2 Nozzle Change Reqd FB1[294].3'; 9412 '~S001R07CN.I.Slr2CycleInterrupted - Seal Cntrl2 Cycle Interrupted FB1[294].4'; 9413 '~S001R07CN.I.Stdw2Flt - Stud Weld 2 Weld Fault FB1[294].5'; 9414 '~S001R07CN.I.Stdw2DlyExcdd - Stud Weld 2 Time Delay Exceeded Flt FB1[294].6'; 9415 '~S001R07CN.I.Stdw2Maint Reqd - Stud Weld 2 Maintenance Required FB1[294].7'; 9416 '~S001R07CN.I.Stdw2Reject - Stud Weld 2 art Reject Fault FB1[294].8'; 9417 '~S001R07CN.I.Rvt2Flt - Rivet Controller 2 Fault FB1[294].9'; 9418 '~S001R07CN.I.Rvt2DlyExcdd - Rivet Cntrl 2 Time Delay Exceeded Flt FB1[294].10'; 9419 '~S001R07CN.I.AutoPulledTipByp2 - Auto Pulled Tip Bypass 2 FB1[294].11'; 9420 '~S001R07CN.I.StdWld2EquipmentFlt - Stud Weld 2 Equipment Fault FB1[294].12'; 9421 '~S001R07CN.I.StdWld2BrcktNotPresent - Stud Weld 2 Bracket Not Pres FB1[294].13'; 9422 '~S001R07CN.Ix.LsrWldMntrFlt - Seam Geometry/Laser Weld Monitor Flt FB1[294].14'; 9423 '~S001R07CN.Ix.LsrHeadFlt - Laser Head Fault FB1[294].15'; 9424 '~S001R07CN.Ix.LsrGlsFlt - Glass Fault FB1[294].16'; 9425 '~S001R07CN.Ix.LsrWhlFlt - Pressure Wheel Not In Range Fault FB1[294].17'; 9426 '~S001R07CN.Ix.LsrGeoFlt - Seam Geometry/Laser Bad Process Geo Flt FB1[294].18'; 9427 '~S001R07CN.Ix.LsrHdCollFlt - Laser Head Collision Fault FB1[294].19'; 9428 '~S001R07CN.Ix.LsrHdSysFlt - Laser Head System Fault FB1[294].20'; 9429 '~S001R07CN.Ix.LsrHdFar - Laser Head Far Fault FB1[294].21'; 9430 '~S001R07CN.Ix.LsrHdSftCollFlt - Laser Head Software Collision Flt FB1[294].22'; 9431 '~S001R07CN.I.O.TipChngReqd2 - Weld Cntrl 2 Tip Change Required FB1[294].23'; 9432 '~S001R07CN.I.M.NutDetectFlt2 - Nut Welder 2 Nut Detection Fault FB1[294].24'; 9433 '~S001R07CN.I.M.NutProjFlt2 - Nut Welder 2 Weld Not In Tolerance FB1[294].25'; 9434 '~S001R07CN.I.TCWrongToolInStand - Tool Changer Wrong Tool In Stand FB1[294].26'; 9435 '~Spare FB1[294].27'; 9436 '~Spare FB1[294].28'; 9437 '~Spare FB1[294].29'; 9438 '~Spare FB1[294].30'; 9439 '~Spare FB1[294].31'; 9440 '~S001R07CN.I.VisionCommOK - Vision System Comm Fault FB1[295].0'; 9441 '~S001R07CN.I.OutOfTolerance - Vision System Out Of Tolerance FB1[295].1'; 9442 '~S001R07CN.I.MeasureReject - Vision System Measure Reject FB1[295].2'; 9443 '~S001R07CN.I.VisionSysCalibrationFlt - Vision System Calibration Flt FB1[295].3'; 9444 '~S001R07CN.I.VisionSysFlt - Vision System Flt FB1[295].4'; 9445 '~Spare FB1[295].5'; 9446 '~Spare FB1[295].6'; 9447 '~Spare FB1[295].7'; 9448 '~Spare FB1[295].8'; 9449 '~Spare FB1[295].9'; 9450 '~Spare FB1[295].10'; 9451 '~Spare FB1[295].11'; 9452 '~Spare FB1[295].12'; 9453 '~Spare FB1[295].13'; 9454 '~Spare FB1[295].14'; 9455 '~Spare FB1[295].15'; 9456 '~Spare FB1[295].16'; 9457 '~Spare FB1[295].17'; 9458 '~S001R07CN.M.InteruptCyc - Laser Cyc Interupt Cut Wire And Reject Car FB1[295].18'; 9459 '~S001R07CN.M.SuspectPart Inspect Vehicle And Accept Or Reject FB1[295].19'; 9460 '~S001R07 Power Meter High Power Fault Detected FB1[295].20'; 9461 '~S001R07 Power Meter Low Power Fault Detected FB1[295].21'; 9462 '~Spare FB1[295].22'; 9463 '~Spare FB1[295].23'; 9464 '~Spare FB1[295].24'; 9465 '~Spare FB1[295].25'; 9466 '~Spare FB1[295].26'; 9467 '~Spare FB1[295].27'; 9468 '~Spare FB1[295].28'; 9469 '~Spare FB1[295].29'; 9470 '~Spare FB1[295].30'; 9471 '~Spare FB1[295].31'; 9472 '~Spare FB1[296].0'; 9473 '~Spare FB1[296].1'; 9474 '~Spare FB1[296].2'; 9475 '~Spare FB1[296].3'; 9476 '~Spare FB1[296].4'; 9477 '~Spare FB1[296].5'; 9478 '~Spare FB1[296].6'; 9479 '~Spare FB1[296].7'; 9480 '~Spare FB1[296].8'; 9481 '~Spare FB1[296].9'; 9482 '~Spare FB1[296].10'; 9483 '~Spare FB1[296].11'; 9484 '~Spare FB1[296].12'; 9485 '~Spare FB1[296].13'; 9486 '~Spare FB1[296].14'; 9487 '~Spare FB1[296].15'; 9488 '~Spare FB1[296].16'; 9489 '~Spare FB1[296].17'; 9490 '~Spare FB1[296].18'; 9491 '~Spare FB1[296].19'; 9492 '~Spare FB1[296].20'; 9493 '~Spare FB1[296].21'; 9494 '~Spare FB1[296].22'; 9495 '~Spare FB1[296].23'; 9496 '~Spare FB1[296].24'; 9497 '~Spare FB1[296].25'; 9498 '~Spare FB1[296].26'; 9499 '~Spare FB1[296].27'; 9500 '~Spare FB1[296].28'; 9501 '~Spare FB1[296].29'; 9502 '~Spare FB1[296].30'; 9503 '~Spare FB1[296].31'; 9504 '~Spare FB1[297].0'; 9505 '~Spare FB1[297].1'; 9506 '~Spare FB1[297].2'; 9507 '~Spare FB1[297].3'; 9508 '~Spare FB1[297].4'; 9509 '~Spare FB1[297].5'; 9510 '~Spare FB1[297].6'; 9511 '~Spare FB1[297].7'; 9512 '~Spare FB1[297].8'; 9513 '~Spare FB1[297].9'; 9514 '~Spare FB1[297].10'; 9515 '~Spare FB1[297].11'; 9516 '~Spare FB1[297].12'; 9517 '~Spare FB1[297].13'; 9518 '~Spare FB1[297].14'; 9519 '~Spare FB1[297].15'; 9520 '~Spare FB1[297].16'; 9521 '~Spare FB1[297].17'; 9522 '~Spare FB1[297].18'; 9523 '~Spare FB1[297].19'; 9524 '~Spare FB1[297].20'; 9525 '~Spare FB1[297].21'; 9526 '~Spare FB1[297].22'; 9527 '~Spare FB1[297].23'; 9528 '~Spare FB1[297].24'; 9529 '~Spare FB1[297].25'; 9530 '~Spare FB1[297].26'; 9531 '~Spare FB1[297].27'; 9532 '~Spare FB1[297].28'; 9533 '~Spare FB1[297].29'; 9534 '~Spare FB1[297].30'; 9535 '~Spare FB1[297].31'; 9536 '~Spare FB1[298].0'; 9537 '~Spare FB1[298].1'; 9538 '~Spare FB1[298].2'; 9539 '~Spare FB1[298].3'; 9540 '~Spare FB1[298].4'; 9541 '~Spare FB1[298].5'; 9542 '~Spare FB1[298].6'; 9543 '~Spare FB1[298].7'; 9544 '~Spare FB1[298].8'; 9545 '~Spare FB1[298].9'; 9546 '~Spare FB1[298].10'; 9547 '~Spare FB1[298].11'; 9548 '~Spare FB1[298].12'; 9549 '~Spare FB1[298].13'; 9550 '~Spare FB1[298].14'; 9551 '~Spare FB1[298].15'; 9552 '~Spare FB1[298].16'; 9553 '~Spare FB1[298].17'; 9554 '~Spare FB1[298].18'; 9555 '~Spare FB1[298].19'; 9556 '~Spare FB1[298].20'; 9557 '~Spare FB1[298].21'; 9558 '~Spare FB1[298].22'; 9559 '~Spare FB1[298].23'; 9560 '~Spare FB1[298].24'; 9561 '~Spare FB1[298].25'; 9562 '~Spare FB1[298].26'; 9563 '~Spare FB1[298].27'; 9564 '~Spare FB1[298].28'; 9565 '~Spare FB1[298].29'; 9566 '~Spare FB1[298].30'; 9567 '~Spare FB1[298].31'; 9568 '~Spare FB1[299].0'; 9569 '~Spare FB1[299].1'; 9570 '~Spare FB1[299].2'; 9571 '~Spare FB1[299].3'; 9572 '~Spare FB1[299].4'; 9573 '~Spare FB1[299].5'; 9574 '~Spare FB1[299].6'; 9575 '~Spare FB1[299].7'; 9576 '~Spare FB1[299].8'; 9577 '~Spare FB1[299].9'; 9578 '~Spare FB1[299].10'; 9579 '~Spare FB1[299].11'; 9580 '~Spare FB1[299].12'; 9581 '~Spare FB1[299].13'; 9582 '~Spare FB1[299].14'; 9583 '~Spare FB1[299].15'; 9584 '~Spare FB1[299].16'; 9585 '~Spare FB1[299].17'; 9586 '~Spare FB1[299].18'; 9587 '~Spare FB1[299].19'; 9588 '~Spare FB1[299].20'; 9589 '~Spare FB1[299].21'; 9590 '~Spare FB1[299].22'; 9591 '~Spare FB1[299].23'; 9592 '~Spare FB1[299].24'; 9593 '~Spare FB1[299].25'; 9594 '~Spare FB1[299].26'; 9595 '~Spare FB1[299].27'; 9596 '~Spare FB1[299].28'; 9597 '~Spare FB1[299].29'; 9598 '~Spare FB1[299].30'; 9599 '~Spare FB1[299].31'; 9600 '~S001R08CN.I.RbtCtrlFlt - Control Fault FB1[300].0'; 9601 '~S001R08CN.I.CollDetect - Collision Detect FB1[300].1'; 9602 '~S001R08CN.Ix.RbtPromptBox - View Prompt Box at Teach Pendant FB1[300].2'; 9603 '~Spare FB1[300].3'; 9604 '~Spare FB1[300].4'; 9605 '~Spare FB1[300].5'; 9606 '~Spare FB1[300].6'; 9607 '~Spare FB1[300].7'; 9608 '~Spare FB1[300].8'; 9609 '~Spare FB1[300].9'; 9610 '~Spare FB1[300].10'; 9611 '~S001R08CN.I.Wc1WldFlt -Weld Controller 1 Weld Fault FB1[300].11'; 9612 '~S001R08CN.I.Wc1Flt - Weld Timer Flt - Depress Man Weld To Continue FB1[300].12'; 9613 '~S001R08CN.I.Wc1SGunFlt - Weld Controller 1 Servo Gun Fault FB1[300].13'; 9614 '~S001R08CN.I.Wc1SGunMtrTempFlt - Cntrl 1 Servo Gun Motor Over Temp FB1[300].14'; 9615 '~S001R08CN.I.Td1MtrFlt - Tip Dress 1 Motor Fault FB1[300].15'; 9616 '~S001R08CN.I.WC1XfmrTempFlt - Weld Cntrl 1 Transformer Over Temp FB1[300].16'; 9617 '~S001R08CN.I.AutoTipChng1Flt - Auto Tip Changer 1 Fault FB1[300].17'; 9618 '~S001R08CN.I.Slr1NotReady - Seal Controller 1 Not Ready FB1[300].18'; 9619 '~S001R08CN.I.Slr1MajorFlt - Seal Controller 1 Major Fault FB1[300].19'; 9620 '~S001R08CN.I.Slr1VolNotOk - Seal Controller 1 Volume Not Ok Fault FB1[300].20'; 9621 '~S001R08CN.I.Slr1PurgeFlt - Seal Controller 1 Purge Fault FB1[300].21'; 9622 '~S001R08CN.I.Slr1DoserNot Filled - Seal Cntrl 1 Doser Not Filled FB1[300].22'; 9623 '~S001R08CN.I.Slr1No2ClnMxr - Seal Cntrl1 No 2C In Mixer Fault FB1[300].23'; 9624 '~S001R08CN.I.Slr1NzlBroken - Seal Controller 1 Nozzle Broken Fault FB1[300].24'; 9625 '~S001R08CN.I.Slr1NozzleChgReq - Seal Cntrl1 Nozzle Change Reqd FB1[300].25'; 9626 '~S001R08CN.I.Slr1CycleInterrupted - Seal Cntrl1 Cycle Interrupted FB1[300].26'; 9627 '~S001R08CN.I.Stdw1Flt - Stud Weld 1 Weld Fault FB1[300].27'; 9628 '~S001R08CN.I.Stdw1DlyExcdd - Stud Weld 1 Time Delay Exceeded Flt FB1[300].28'; 9629 '~S001R08CN.I.Stdw1Maint Reqd - Stud Weld 1 Maintenance Required FB1[300].29'; 9630 '~S001R08CN.I.Stdw1Reject - Stud Weld 1 art Reject Fault FB1[300].30'; 9631 '~S001R08CN.I.Rvt1Flt - Rivet Controller 1 Fault FB1[300].31'; 9632 '~S001R08CN.I.Rvt1DlyExcdd - Rivet Cntrl 1 Time Delay Exceeded Flt FB1[301].0'; 9633 '~S001R08CN.I.AutoPulledTipByp1 - Auto Pulled Tip Bypass 1 FB1[301].1'; 9634 '~S001R08CN.I.StdWld1EquipmentFlt - Stud Weld 1 Equipment Fault FB1[301].2'; 9635 '~S001R08CN.I.StdWld1BrcktNotPresent - Stud Weld 1 Bracket Not Pres FB1[301].3'; 9636 '~S001R08CN.I.PierceFlt - Pierce Fault FB1[301].4'; 9637 '~S001R08CN.I.NoVisionMeasErr - Vision System Measurement Error FB1[301].5'; 9638 '~S001R08CN.I.VisionSysCalErr - Vision System Calibration Fault FB1[301].6'; 9639 '~S001R08CN.I.VisionSysErr - Vision System Error FB1[301].7'; 9640 '~S001R08CN.I.RackOutOfTolerance - Vision Sys Rack Out Of Tolerance FB1[301].8'; 9641 '~S001R08CN.Ix.TorqFlt - Torque Not Ok FB1[301].9'; 9642 '~S001R08CN.Ix.MwFlt - Mig Weld Controller Fault FB1[301].10'; 9643 '~S001R08CN.Ix.MwWireStuckFlt - Mig Welder Wire Stuck FB1[301].11'; 9644 '~S001R08CN.Ix.MwWldFlt - Mig Welder Bad Bronze Weld Indicator Flt FB1[301].12'; 9645 '~S001R08CN.I.O.TipChngReqd1 - Weld Cntrl 1 Tip Change Required FB1[301].13'; 9646 '~S001R08CN.I.M.NutDetectFlt1 - Nut Welder 1 Nut Detection Fault FB1[301].14'; 9647 '~S001R08CN.I.M.NutProjFlt1 - Nut Welder 1 Weld Not In Tolerance FB1[301].15'; 9648 '~S001R08CN.M.WrongRivetAtNose - Remove Wrong Rivet At Nose FB1[301].16'; 9649 '~S001R08CN.Ix.MwWldLimitErr - Mig Welder CurrentVoltage Out of Tolerance FB1[301].17'; 9650 '~S001R08CN.Ix.MigRdy Mig Welder Not Ready FB1[301].18'; 9651 '~Spare FB1[301].19'; 9652 '~Spare FB1[301].20'; 9653 '~S001R08CN.I.Wc2WldFlt -Weld Controller 2 Weld Fault FB1[301].21'; 9654 '~S001R08CN.I.Wc2Flt - Weld Timer 